       ELSIF "DB110_Interf_Program_M1".Status_IF[16].IF_is_on_1_Position AND "DB123_MH_IO_Signals".MH[16].IN.MH_Manual_Mode AND
           (#TempStationNo > 0 AND #TempStationNo < 101) THEN
           "DB619_State_MPart".ToolMa[#TmpMachineNumber].ToolNo := "DB941_Tool_alloc_manual_MH".MH[16].Alloc_stationTool[#TempStationNo];
       ELSE
           "DB619_State_MPart".ToolMa[#TmpMachineNumber].ToolNo := "DB940_Tool_alloc_automatic".Alloc_stationTool[#TempStationNo];
       END_IF;

       "DB619_State_MPart".ToolMa[#TmpMachineNumber].StationActive := True;
       "DB619_State_MPart".ToolMa[#TmpMachineNumber].StationNo := INT_TO_BYTE(#TempStationNo);
   END_IF;

   #TmpActToolNo := "DB619_State_MPart".ToolMa[#TmpMachineNumber].ToolNo;

   //-----------------------------------------------------------------
   // Check if tool no. between 1 and Amount tools if OK get data
   // ----------------------------------------------------------------
   IF (#TmpActToolNo > 0 AND
       #TmpActToolNo < "AmountTools") AND
      #IO_PartShotNoNew =  0 
    THEN
         #IO_PartShotNoNew:=  1;
         // Get tool values                                               
         "DB619_State_MPart".ToolMa[#TmpMachineNumber].Tool:= "DB930_Tools".Tool[#TmpActToolNo];
         // Get shot values; 
         IF (#TmpActToolNo > 0 AND
             #TmpActToolNo <= "AmountToolsDB")
         THEN
             "DB619_State_MPart".ShotMa[#TmpMachineNumber].Tool := "DB925_ShotData_1".Tool[#TmpActToolNo];

         ELSIF (#TmpActToolNo > "AmountToolsDB" AND #TmpActToolNo <= (2*"AmountToolsDB")) THEN
             "DB619_State_MPart".ShotMa[#TmpMachineNumber].Tool := "DB926_ShotData_2".Tool[#TmpActToolNo-"AmountToolsDB"];
         END_IF;

     ELSIF NOT (#TmpActToolNo > 0 AND #TmpActToolNo < "AmountToolsDB") THEN
         // Fault wrong tool no.    
         IF NOT #IO_Faults.FLT_WrongToolNumber AND
             "DB619_State_MPart".ToolMa[#TmpMachineNumber].StationActive AND
             NOT "DB619_State_MPart".ToolMa[#TmpMachineNumber].StationFinished THEN
               #IO_Faults.FLT_WrongToolNumber  := True;
               #IO_NewFault := True;
         END_IF;  
     END_IF;

   //-----------------------------------------------------------------------------------------
   // Check if new Tool is deselected 
   // ----------------------------------------------------------------------------------------
     IF NOT "DB619_State_MPart".ToolMa[#TmpMachineNumber].Tool.EnableTool AND
         "DB619_State_MPart".ToolMa[#TmpMachineNumber].StationActive THEN
         "DB619_State_MPart".ToolMa[#TmpMachineNumber].StationFinished := TRUE;
         "DB619_State_MPart".ToolMa[#TmpMachineNumber].ShotFound := FALSE;
         "DB619_State_MPart".ToolMa[#TmpMachineNumber].ToolNo := 0;
         "DB619_State_MPart".ToolMa[#TmpMachineNumber].PartShot := 0;
         "DB619_State_MPart".ShotMa[#TmpMachineNumber].ShotData.MH_No := 0;

         #IO_Faults.Reserve3 := TRUE;
   END_IF;


   //-----------------------------------------------------------------------------------------
   // Check if new partshot no. exist than get new MH no. and Shotvalues and set ShoFound 
   // ----------------------------------------------------------------------------------------
   IF #IO_PartShotNoNew <> "DB619_State_MPart".ToolMa[#TmpMachineNumber].PartShot AND
       "DB619_State_MPart".ToolMa[#TmpMachineNumber].StationActive
        THEN
            "DB619_State_MPart".ToolMa[#TmpMachineNumber].PartShot := #IO_PartShotNoNew;

         // Get mixinghead no. of selected part shot
            IF (#TmpActToolNo > 0 AND #TmpActToolNo < "AmountToolsDB") THEN
                #MH_No := "DB925_ShotData_1".Tool[#TmpActToolNo].Shot[#IO_PartShotNoNew].MHNo;
            ELSIF (#TmpActToolNo > "AmountToolsDB" AND #TmpActToolNo <= (2*"AmountToolsDB")) THEN
                #MH_No := "DB926_ShotData_2".Tool[#TmpActToolNo-"AmountToolsDB"].Shot[#IO_PartShotNoNew].MHNo;
            END_IF;

         "DB619_State_MPart".ShotMa[#TmpMachineNumber].ShotData.MH_No := INT_TO_BYTE(#MH_No);
             // Check mixinghead no. between 1 and 12
             IF #MH_No > 0 AND #MH_No < 13 THEN
                   // Mixinghead is connected at this machine
                   #MHNoShift := 1;
                   #MHNoBinary := SHL(IN :=  #MHNoShift, N := #MH_No -1);
                   #TmpMHatThisMachine := ("DB700_Machine".Machine[#TmpMachineNumber].MH_at_Machine AND #MHNoBinary) <> 0;
             ELSE
                   // Fault wrong mixinghead no. 
                 IF NOT  #IO_Faults.FLT_WrongMixingheadNumber AND "DB619_State_MPart".ToolMa[#TmpMachineNumber].StationActive THEN    // Must be wrong mixinghead no.                                                  
                     #IO_Faults.FLT_WrongMixingheadNumber := True;
                     #IO_Faults.FLT_WrongMixingheadNumber := False;
                     // #IO_NewFault := True;
                     //"DB619_State_MPart".ToolMa[#TmpMachineNumber].StationActive := FALSE;
                     //"DB619_State_MPart".ToolMa[#TmpMachineNumber].StationFinished := TRUE;
                 END_IF;
             END_IF;

   // Get shot values of current foamingcycle
             "DB619_State_MPart".ShotMa[#TmpMachineNumber].ShotData.ShotDisabled := "DB619_State_MPart".ShotMa[#TmpMachineNumber].Tool.Shot[#IO_PartShotNoNew].PartShotDisable;
             "DB619_State_MPart".ShotMa[#TmpMachineNumber].ShotData.CP_AfterShot := "DB619_State_MPart".ShotMa[#TmpMachineNumber].Tool.Shot[#IO_PartShotNoNew].CPMoveAfterShot;
             "DB619_State_MPart".ShotMa[#TmpMachineNumber].ShotData.Foamingtime := "DB619_State_MPart".ShotMa[#TmpMachineNumber].Tool.Shot[#IO_PartShotNoNew].FoamingTime;
             "DB619_State_MPart".ShotMa[#TmpMachineNumber].ShotData.PurgeMH_AfterShot := "DB619_State_MPart".ShotMa[#TmpMachineNumber].Tool.Shot[#IO_PartShotNoNew].PurgeMHAfterShot;

             "DB619_State_MPart".ShotMa[#TmpMachineNumber].ShotData.Flow[1] := "DB619_State_MPart".ShotMa[#TmpMachineNumber].Tool.Shot[#IO_PartShotNoNew].Flow[1];
             "DB619_State_MPart".ShotMa[#TmpMachineNumber].ShotData.Flow[2] := "DB619_State_MPart".ShotMa[#TmpMachineNumber].Tool.Shot[#IO_PartShotNoNew].Flow[2];
             "DB619_State_MPart".ShotMa[#TmpMachineNumber].ShotData.Flow[3] := "DB619_State_MPart".ShotMa[#TmpMachineNumber].Tool.Shot[#IO_PartShotNoNew].Flow[3];
             "DB619_State_MPart".ShotMa[#TmpMachineNumber].ShotData.Flow[4] := "DB619_State_MPart".ShotMa[#TmpMachineNumber].Tool.Shot[#IO_PartShotNoNew].Flow[4];
             "DB619_State_MPart".ShotMa[#TmpMachineNumber].ShotData.Flow[5] := "DB619_State_MPart".ShotMa[#TmpMachineNumber].Tool.Shot[#IO_PartShotNoNew].Flow[5];
             "DB619_State_MPart".ShotMa[#TmpMachineNumber].ShotData.Flow[6] := "DB619_State_MPart".ShotMa[#TmpMachineNumber].Tool.Shot[#IO_PartShotNoNew].Flow[6];
             "DB619_State_MPart".ShotMa[#TmpMachineNumber].ShotData.Pressure[1] := "DB619_State_MPart".ShotMa[#TmpMachineNumber].Tool.Shot[#IO_PartShotNoNew].Pressure[1];
             "DB619_State_MPart".ShotMa[#TmpMachineNumber].ShotData.Pressure[2] := "DB619_State_MPart".ShotMa[#TmpMachineNumber].Tool.Shot[#IO_PartShotNoNew].Pressure[2];
             "DB619_State_MPart".ShotMa[#TmpMachineNumber].ShotData.Pressure[3] := "DB619_State_MPart".ShotMa[#TmpMachineNumber].Tool.Shot[#IO_PartShotNoNew].Pressure[3];
             "DB619_State_MPart".ShotMa[#TmpMachineNumber].ShotData.Pressure[4] := "DB619_State_MPart".ShotMa[#TmpMachineNumber].Tool.Shot[#IO_PartShotNoNew].Pressure[4];
             "DB619_State_MPart".ShotMa[#TmpMachineNumber].ShotData.Pressure[5] := "DB619_State_MPart".ShotMa[#TmpMachineNumber].Tool.Shot[#IO_PartShotNoNew].Pressure[5];
             "DB619_State_MPart".ShotMa[#TmpMachineNumber].ShotData.Pressure[6] := "DB619_State_MPart".ShotMa[#TmpMachineNumber].Tool.Shot[#IO_PartShotNoNew].Pressure[6];

             "DB619_State_MPart".ShotMa[#TmpMachineNumber].ShotData."2PointAdjustment"[1] := "DB619_State_MPart".ShotMa[#TmpMachineNumber].Tool.Shot[#IO_PartShotNoNew]."2PoinMovement_Comp01";
             "DB619_State_MPart".ShotMa[#TmpMachineNumber].ShotData."2PointAdjustment"[2] := "DB619_State_MPart".ShotMa[#TmpMachineNumber].Tool.Shot[#IO_PartShotNoNew]."2PoinMovement_Comp02";
             "DB619_State_MPart".ShotMa[#TmpMachineNumber].ShotData."2PointAdjustment"[3] := "DB619_State_MPart".ShotMa[#TmpMachineNumber].Tool.Shot[#IO_PartShotNoNew]."2PoinMovement_Comp03";
             "DB619_State_MPart".ShotMa[#TmpMachineNumber].ShotData."2PointAdjustment"[4] := "DB619_State_MPart".ShotMa[#TmpMachineNumber].Tool.Shot[#IO_PartShotNoNew]."2PoinMovement_Comp04";
             "DB619_State_MPart".ShotMa[#TmpMachineNumber].ShotData."2PointAdjustment"[5] := "DB619_State_MPart".ShotMa[#TmpMachineNumber].Tool.Shot[#IO_PartShotNoNew]."2PoinMovement_Comp05";
             "DB619_State_MPart".ShotMa[#TmpMachineNumber].ShotData."2PointAdjustment"[6] := "DB619_State_MPart".ShotMa[#TmpMachineNumber].Tool.Shot[#IO_PartShotNoNew]."2PoinMovement_Comp06";

             "DB619_State_MPart".ShotMa[#TmpMachineNumber].ShotData.PartCounter := "DB619_State_MPart".ShotMa[#TmpMachineNumber].Tool.Shot[#IO_PartShotNoNew].PartCounter;


             "DB606_PV_Machine".Machine[#TmpMachineNumber].ShotTime.PV_SetV.Value := "DB619_State_MPart".ShotMa[#TmpMachineNumber].Tool.Shot[#IO_PartShotNoNew].FoamingTime;

   // Fault at tool is active      
   #IO_FaultAtStation := #IO_Faults.FLT_WrongToolNumber       OR
                         #IO_Faults.FLT_WrongMixingheadNumber OR
                         #IO_Faults.FLT_NewNoTooEarly;

   // Set shot found if tool is enabled                      
                         IF "DB619_State_MPart".ToolMa[#TmpMachineNumber].StationActive  AND NOT
                                              #IO_FaultAtStation  AND
                                              #IN_EnableTool      AND
                                              #TmpMHatThisMachine AND
                                              "DB619_State_MPart".ToolMa[#TmpMachineNumber].Tool.EnableTool
      THEN            
          "DB619_State_MPart".ToolMa[#TmpMachineNumber].ShotFound := True;
      ELSE       
          "DB619_State_MPart".ToolMa[#TmpMachineNumber].ShotFound := FALSE;
      END_IF;
    END_IF;

   //------------------------------------------------------------------------------------------
   // New Partshot no. -> Shotend, Shotbreak, next shot at this machine
   // -----------------------------------------------------------------------------------------
    IF  ("DB619_State_MPart".ToolMa[#TmpMachineNumber].StationActive AND NOT
        "DB619_State_MPart".ToolMa[#TmpMachineNumber].ShotFound)     OR
        "DB619_State_MPart".Cycle[#TmpMachineNumber].PulsShotend
       THEN  
           IF "DB619_State_MPart".ToolMa[#TmpMachineNumber].PartShot <= BYTE_TO_INT("DB619_State_MPart".ToolMa[#TmpMachineNumber].Tool.PartShot_Amount) THEN
               #IO_PartShotNoNew := "DB619_State_MPart".ToolMa[#TmpMachineNumber].PartShot + 1;
               "DB619_State_MPart".ToolMa[#TmpMachineNumber].ShotFound := FALSE;
           END_IF;

       END_IF;

       // Station finished: shots done; cycle stopped; fault level 1; station no. = 0
       IF "DB619_State_MPart".ToolMa[#TmpMachineNumber].PartShot > BYTE_TO_INT("DB619_State_MPart".ToolMa[#TmpMachineNumber].Tool.PartShot_Amount) OR
          "DB009_Faults".Fault_State_Grp_1_M1                 OR
          "DB619_State_MPart".ToolMa[#TmpMachineNumber].StopCycle
       THEN
           "DB619_State_MPart".ToolMa[#TmpMachineNumber].StationFinished := TRUE;
           "DB619_State_MPart".ToolMa[#TmpMachineNumber].ShotFound := FALSE;
           "DB619_State_MPart".ToolMa[#TmpMachineNumber].ToolNo := 0;
           "DB619_State_MPart".ToolMa[#TmpMachineNumber].PartShot := 0;
           "DB619_State_MPart".ShotMa[#TmpMachineNumber].ShotData.MH_No := 0;
       END_IF;

       IF  #IO_Faults.FLT_WrongToolNumber       OR
           #IO_Faults.FLT_WrongMixingheadNumber OR
           #IO_Faults.FLT_NewNoTooEarly         OR
           #IO_Faults.Reserve3
         THEN
           #IO_FaultLevel_1 := TRUE;
       END_IF;
END_FUNCTION_BLOCK

FUNCTION_BLOCK "FB1931_ToolAllocationList"   // FB1931, SCL
{ S7_Optimized_Access := 'TRUE' }
VERSION : 0.1
   VAR
      Alloc_stationTool : Array[0..30] of Int;
      SaveSortProgs : Array[0..20] of Int;
   END_VAR
   VAR_TEMP
      j : Int;
      i : Int;
      z : Int;
      TiLoop : Int;
      TiLoopSave : Int;
      TiLoopMH : Int;
      Ti_alloc_list : Int;
      Amount_tools : Int;
      MH_No_hand_allocation : Int;
      Offset_SavedProgsList : Int;
      Offset_AllocateList : Int;
      LimitSavedProgList : Int;
      Amount_Saved_tools : Int;
      tool_okay : Bool;
   END_VAR
   // Alloc_stationTool[0] := 0;
   // Alloc_stationTool[1] := 0;
   // Alloc_stationTool[2] := 0;
   // Alloc_stationTool[3] := 0;
   // Alloc_stationTool[4] := 0;
   // Alloc_stationTool[5] := 0;
   // Alloc_stationTool[6] := 0;
   // Alloc_stationTool[7] := 0;
   // Alloc_stationTool[8] := 0;
   // Alloc_stationTool[9] := 0;
   // Alloc_stationTool[10] := 0;
   // Alloc_stationTool[11] := 0;
   // Alloc_stationTool[12] := 0;
   // Alloc_stationTool[13] := 0;
   // Alloc_stationTool[14] := 0;
   // Alloc_stationTool[15] := 0;
   // Alloc_stationTool[16] := 0;
   // Alloc_stationTool[17] := 0;
   // Alloc_stationTool[18] := 0;
   // Alloc_stationTool[19] := 0;
   // Alloc_stationTool[20] := 0;
   // Alloc_stationTool[21] := 0;
   // Alloc_stationTool[22] := 0;
   // Alloc_stationTool[23] := 0;
   // Alloc_stationTool[24] := 0;
   // Alloc_stationTool[25] := 0;
   // Alloc_stationTool[26] := 0;
   // Alloc_stationTool[27] := 0;
   // Alloc_stationTool[28] := 0;
   // Alloc_stationTool[29] := 0;
   // Alloc_stationTool[30] := 0;
BEGIN
   // Limit values

   "DB939_Tool_alloc_HMI".Selected_prog := LIMIT(MN := 1, IN := "DB939_Tool_alloc_HMI".Selected_prog, MX := 30);
   "DB939_Tool_alloc_HMI".Selected_SavedProg := LIMIT(MN := 0, IN := "DB939_Tool_alloc_HMI".Selected_SavedProg, MX := 20);
   "DB939_Tool_alloc_HMI".Limit_allocation_list := LIMIT(MN := 1, IN := "DB939_Tool_alloc_HMI".Limit_allocation_list, MX := 30);

   FOR #TiLoop := 0 TO 30 DO
       "DB939_Tool_alloc_HMI".Alloc_stationTool[#TiLoop] := LIMIT(MN := 0, IN := "DB939_Tool_alloc_HMI".Alloc_stationTool[#TiLoop], MX := "AmountTools");
   END_FOR;

   REGION Select manual/auto
       // Switch for choosing manual or automatic allocation on the Screen "ProgramAllocation"  
       IF "DB939_Tool_alloc_HMI".Select_hand_automatic_alloc = TRUE THEN
           "DB939_Tool_alloc_HMI".Tool_allocation_automatic := FALSE;
           "DB939_Tool_alloc_HMI".Tool_allocation_manual := TRUE;
       ELSE
           "DB939_Tool_alloc_HMI".Tool_allocation_automatic := TRUE;
           "DB939_Tool_alloc_HMI".Tool_allocation_manual := FALSE;
       END_IF;
   END_REGION

   // Current selected mixing head number for Hand allocation
   #MH_No_hand_allocation := "DB939_Tool_alloc_HMI".MH_No_selected;

   REGION Visibility MH arrows 
       // Visibility of arrow for decreasing Mixing head number
       IF "DB939_Tool_alloc_HMI".Tool_allocation_manual = TRUE AND #MH_No_hand_allocation > 1 THEN
           "DB939_Tool_alloc_HMI".MH_Nr_decrease_visible := TRUE;
       ELSE
           "DB939_Tool_alloc_HMI".MH_Nr_decrease_visible := FALSE;
       END_IF;

       // Visibility of arrow for increasing Mixing head number
       IF "DB939_Tool_alloc_HMI".Tool_allocation_manual = TRUE AND #MH_No_hand_allocation < "DB790_PlantParameter".AmountMH THEN
           "DB939_Tool_alloc_HMI".MH_Nr_increase_visible := TRUE;
       ELSE
           "DB939_Tool_alloc_HMI".MH_Nr_increase_visible := FALSE;
       END_IF;
   END_REGION

   REGION Page AllocationList
       // Depending on amound of manual programs limit list and pages
       IF "DB704_MH_Value".Mixinghead[#MH_No_hand_allocation].With99program = FALSE AND "DB939_Tool_alloc_HMI".Tool_allocation_automatic = FALSE THEN
           "DB939_Tool_alloc_HMI".Limit_allocation_page := 1;
           "DB939_Tool_alloc_HMI".Limit_allocation_list := 9;
       ELSIF "DB704_MH_Value".Mixinghead[#MH_No_hand_allocation].With99program = TRUE AND "DB939_Tool_alloc_HMI".Tool_allocation_automatic = FALSE THEN
           "DB939_Tool_alloc_HMI".Limit_allocation_page := 4;
           IF "DB939_Tool_alloc_HMI".AllocList_page >= 4 THEN
               "DB939_Tool_alloc_HMI".Limit_allocation_list := 9;
           ELSE
               "DB939_Tool_alloc_HMI".Limit_allocation_list := 30;
           END_IF;
       ELSIF "DB939_Tool_alloc_HMI".Tool_allocation_automatic = TRUE THEN
         //Depending on the amount of the stationsnumber   
           "DB939_Tool_alloc_HMI".Limit_allocation_page := (("DB790_PlantParameter".AmountToolStation -1 ) / (30))+1;
           IF "DB939_Tool_alloc_HMI".AllocList_page = "DB939_Tool_alloc_HMI".Limit_allocation_page  AND ("DB790_PlantParameter".AmountToolStation MOD 30) <> 0 THEN
               "DB939_Tool_alloc_HMI".Limit_allocation_list := ("DB790_PlantParameter".AmountToolStation MOD 30);
           ELSE
               "DB939_Tool_alloc_HMI".Limit_allocation_list := 30;
           END_IF;
       ELSE   
           "DB939_Tool_alloc_HMI".Limit_allocation_page := 7;
           "DB939_Tool_alloc_HMI".Limit_allocation_list := 30;
       END_IF;

       IF "DB939_Tool_alloc_HMI".AllocList_increase THEN
           "DB939_Tool_alloc_HMI".AllocList_page := "DB939_Tool_alloc_HMI".AllocList_page + 1;
           "DB939_Tool_alloc_HMI".AllocList_increase := False;
       ELSIF "DB939_Tool_alloc_HMI".AllocList_decrease THEN
           "DB939_Tool_alloc_HMI".AllocList_page := "DB939_Tool_alloc_HMI".AllocList_page - 1;
           "DB939_Tool_alloc_HMI".AllocList_decrease := False;
       END_IF;
       // Limit
       "DB939_Tool_alloc_HMI".AllocList_page := LIMIT(MN := 1, IN := "DB939_Tool_alloc_HMI".AllocList_page, MX := "DB939_Tool_alloc_HMI".Limit_allocation_page);
       // Create offset
       #Offset_AllocateList := ("DB939_Tool_alloc_HMI".AllocList_page - 1) * 30;
   END_REGION

   REGION Useable Alloc arrows
    // This part is used for if you can alloc the programm to the allocaationlist by yourself 
    // or automatically by the inferface
       IF "DB939_Tool_alloc_HMI".Tool_allocation_automatic = TRUE AND "DB790_PlantParameter".Bit.ProgrammNofromInterface = TRUE THEN
           IF  ("DB790_PlantParameter".AmountMouldCarrier MOD 30) <> 0 THEN
               IF "DB939_Tool_alloc_HMI".AllocList_page = ((("DB790_PlantParameter".AmountMouldCarrier - 1) / 30)+1) THEN
                    "DB939_Tool_alloc_HMI".Operability_selected_line := ("DB790_PlantParameter".AmountMouldCarrier MOD 30);
                ELSIF   "DB939_Tool_alloc_HMI".AllocList_page < ((("DB790_PlantParameter".AmountMouldCarrier - 1) / 30)+1) THEN
                   "DB939_Tool_alloc_HMI".Operability_selected_line := 30;
                ELSE
                   "DB939_Tool_alloc_HMI".Operability_selected_line := 0;
               END_IF;
           ELSE
               IF "DB939_Tool_alloc_HMI".AllocList_page <= ((("DB790_PlantParameter".AmountMouldCarrier - 1) / 30)+1) THEN
                    "DB939_Tool_alloc_HMI".Operability_selected_line := 30;
               ELSE
                   "DB939_Tool_alloc_HMI".Operability_selected_line := 0;
               END_IF;
           END_IF;
       ELSE 
           "DB939_Tool_alloc_HMI".Operability_selected_line := 0;
       END_IF;

       IF "DB939_Tool_alloc_HMI".Selected_prog <= "DB939_Tool_alloc_HMI".Operability_selected_line THEN
           "DB939_Tool_alloc_HMI".Selected_prog := 0;
       END_IF;
   END_REGION
   REGION Visibility Alloc arrows
       IF "DB939_Tool_alloc_HMI".AllocList_page < "DB939_Tool_alloc_HMI".Limit_allocation_page THEN
           "DB939_Tool_alloc_HMI".AllocList_increase_visible := TRUE;
       ELSE    
           "DB939_Tool_alloc_HMI".AllocList_increase_visible := FALSE;
       END_IF;

       IF "DB939_Tool_alloc_HMI".AllocList_page > 1 THEN
           "DB939_Tool_alloc_HMI".AllocList_decrease_visible := TRUE;
       ELSE
           "DB939_Tool_alloc_HMI".AllocList_decrease_visible := FALSE;
       END_IF;
   END_REGION

   REGION Page SavedProgsList
       // Depending on the saved tools. Limit saved list
       #Amount_Saved_tools := 0;
       FOR #TiLoop := 1 TO "AmountTools" DO
           IF "DB933_SaveSortProgs".SaveSortTool[#TiLoop] <> 0 THEN
               #Amount_Saved_tools := #Amount_Saved_tools + 1;
           END_IF;
       END_FOR;
       IF #Amount_Saved_tools > 0 THEN
           #LimitSavedProgList := ((#Amount_Saved_tools - 1) / 20) + 1;
       ELSE
           #LimitSavedProgList := 1;
       END_IF;


       IF "DB939_Tool_alloc_HMI".SavedProgs_increase THEN
           "DB939_Tool_alloc_HMI".SavedProgs_page := "DB939_Tool_alloc_HMI".SavedProgs_page + 1;
           "DB939_Tool_alloc_HMI".SavedProgs_increase := False;
       ELSIF "DB939_Tool_alloc_HMI".SavedProgs_decrease THEN
           "DB939_Tool_alloc_HMI".SavedProgs_page := "DB939_Tool_alloc_HMI".SavedProgs_page - 1;
           "DB939_Tool_alloc_HMI".SavedProgs_decrease := False;
       END_IF;
       // Limit
       "DB939_Tool_alloc_HMI".SavedProgs_page := LIMIT(MN := 1, IN := "DB939_Tool_alloc_HMI".SavedProgs_page, MX := #LimitSavedProgList);
       // Create offset
       #Offset_SavedProgsList := ("DB939_Tool_alloc_HMI".SavedProgs_page - 1) * 20;
   END_REGION

   REGION Visibility SavedProgList arrows
       IF "DB939_Tool_alloc_HMI".SavedProgs_page < #LimitSavedProgList THEN
           "DB939_Tool_alloc_HMI".SavedProgs_increase_visible := TRUE;
       ELSE
           "DB939_Tool_alloc_HMI".SavedProgs_increase_visible := FALSE;
       END_IF;

       IF "DB939_Tool_alloc_HMI".SavedProgs_page > 1 THEN
           "DB939_Tool_alloc_HMI".SavedProgs_decrease_visible := TRUE;
       ELSE
           "DB939_Tool_alloc_HMI".SavedProgs_decrease_visible := FALSE;
       END_IF;
   END_REGION

   REGION Clear SavedProgsList
       FOR #z := 0 TO "AmountTools" DO
           // Clear list
           "DB933_SaveSortProgs".SaveSortTool[#z] := 0;
       END_FOR;
   END_REGION

   REGION Create SavedProgsList
       // Check if part shots available or not for allocation list
       #j := 1;
       FOR #TiLoop := 1 TO "AmountTools" DO
           IF "DB930_Tools".Tool[#TiLoop].PartShot_Amount <> 0 THEN
               "DB933_SaveSortProgs".SaveSortTool[#j] := #TiLoop;
               #j := #j + 1;
           END_IF;
       END_FOR;
   END_REGION

   REGION Copy Part of list savedprogslist to actual HMI
       FOR #TiLoop := 1 TO 20 DO
           "DB939_Tool_alloc_HMI".SaveSortProgs[#TiLoop] := "DB933_SaveSortProgs".SaveSortTool[#TiLoop + #Offset_SavedProgsList];
       END_FOR;
   END_REGION

   REGION Delete selected tool allocation
       IF "DB939_Tool_alloc_HMI".Delete_selected_tool <> 0 THEN
           "DB939_Tool_alloc_HMI".Alloc_stationTool["DB939_Tool_alloc_HMI".Delete_selected_tool] := 0;
           "DB939_Tool_alloc_HMI".Delete_selected_tool := 0;
       END_IF;
   END_REGION

   REGION Delete selected tool from Mould Editor in all allocation lists
       IF "DB939_Tool_alloc_HMI"."Delete_tool_in _all_allocations" AND "DB_MouldEditor_HMI".uData.sStatusBits.xFaultDeleteProgram THEN
           // search tool in automatic allocation list
           FOR #TiLoop := 1 TO "InterfaceVisu".AmountAlloactionAutomatic DO
               IF "DB940_Tool_alloc_automatic".Alloc_stationTool[#TiLoop] = "DB_MouldEditor_HMI".uData.sSelected.iTool THEN
                   "DB940_Tool_alloc_automatic".Alloc_stationTool[#TiLoop] := 0;
               END_IF;
           END_FOR;
           // search tool in all manual allocation lists
           FOR #TiLoopMH := 1 TO "DB790_PlantParameter".AmountMH DO
               IF "DB704_MH_Value".Mixinghead[#TiLoopMH].With99program THEN
                   #Ti_alloc_list := 99;
               ELSE
                   #Ti_alloc_list := 9;
               END_IF;

               FOR #TiLoop := 1 TO #Ti_alloc_list DO
                   IF "DB941_Tool_alloc_manual_MH".MH[#TiLoopMH].Alloc_stationTool[#TiLoop] = "DB_MouldEditor_HMI".uData.sSelected.iTool THEN
                       "DB941_Tool_alloc_manual_MH".MH[#TiLoopMH].Alloc_stationTool[#TiLoop] := 0;
                   END_IF;
               END_FOR;
           END_FOR;
           // reset bits to delete and for PopUp
           "DB939_Tool_alloc_HMI"."Delete_tool_in _all_allocations" := FALSE;
           "DB_MouldEditor_HMI".uData.sStatusBits.xFaultDeleteProgram := FALSE;
           "DB_MouldEditor_HMI".uData.sStatusBits.xDeleteProgram := TRUE; // <-- delete tool
       END_IF;
   END_REGION

   REGION assign saved tool to selected tool    
       IF "DB939_Tool_alloc_HMI".Selected_SavedProg <> 0 THEN
           // If no programm is allocated set new programm
           IF "DB939_Tool_alloc_HMI".Alloc_stationTool["DB939_Tool_alloc_HMI".Selected_prog] = 0 THEN
               "DB939_Tool_alloc_HMI".Alloc_stationTool["DB939_Tool_alloc_HMI".Selected_prog] := "DB933_SaveSortProgs".SaveSortTool["DB939_Tool_alloc_HMI".Selected_SavedProg + #Offset_SavedProgsList];
               "DB939_Tool_alloc_HMI".Selected_SavedProg := 0;
               "DB939_Tool_alloc_HMI".Overwrite_not_allowed := FALSE;
           ELSIF "DB939_Tool_alloc_HMI".Alloc_stationTool["DB939_Tool_alloc_HMI".Selected_prog] = "DB933_SaveSortProgs".SaveSortTool["DB939_Tool_alloc_HMI".Selected_SavedProg + #Offset_SavedProgsList] THEN
               "DB939_Tool_alloc_HMI".Selected_SavedProg := 0;
           ELSE
               "DB939_Tool_alloc_HMI".Overwrite_not_allowed := TRUE;
               IF "DB939_Tool_alloc_HMI".Overwrite_selected_tool = TRUE THEN
                   "DB939_Tool_alloc_HMI".Alloc_stationTool["DB939_Tool_alloc_HMI".Selected_prog] := "DB933_SaveSortProgs".SaveSortTool["DB939_Tool_alloc_HMI".Selected_SavedProg + #Offset_SavedProgsList];
                   "DB939_Tool_alloc_HMI".Selected_SavedProg := 0;
                   "DB939_Tool_alloc_HMI".Overwrite_not_allowed := FALSE;
                   "DB939_Tool_alloc_HMI".Overwrite_selected_tool := FALSE;
               END_IF;
           END_IF;
       ELSE    
           "DB939_Tool_alloc_HMI".Overwrite_not_allowed := FALSE;
       END_IF;
   END_REGION

   REGION Allocationlist number changed
       // If any allocation list no changed, store it to the right DB
       FOR #TiLoop := 1 TO 30 DO
           IF "DB939_Tool_alloc_HMI".Alloc_stationTool[#TiLoop] <> #Alloc_stationTool[#TiLoop] THEN
               IF "DB939_Tool_alloc_HMI".Tool_allocation_automatic = TRUE THEN
                   "DB940_Tool_alloc_automatic".Alloc_stationTool[#TiLoop + #Offset_AllocateList] := "DB939_Tool_alloc_HMI".Alloc_stationTool[#TiLoop];
               ELSE
                   "DB941_Tool_alloc_manual_MH".MH["DB939_Tool_alloc_HMI".MH_No_selected].Alloc_stationTool[#TiLoop + #Offset_AllocateList] := "DB939_Tool_alloc_HMI".Alloc_stationTool[#TiLoop];
               END_IF;
           END_IF;
       END_FOR;
   END_REGION

   REGION Copy Part of allocat list to actual HMI


       FOR #TiLoop := 1 TO 30 DO
           IF "DB939_Tool_alloc_HMI".Tool_allocation_automatic = TRUE THEN
               "DB939_Tool_alloc_HMI".Alloc_stationTool[#TiLoop] := "DB940_Tool_alloc_automatic".Alloc_stationTool[#TiLoop + #Offset_AllocateList];
           ELSE
               "DB939_Tool_alloc_HMI".Alloc_stationTool[#TiLoop] := "DB941_Tool_alloc_manual_MH".MH["DB939_Tool_alloc_HMI".MH_No_selected].Alloc_stationTool[#TiLoop + #Offset_AllocateList];
           END_IF;
           // Depending on BCD switch load 9 or 30 (99) programs in the list
           IF ("DB704_MH_Value".Mixinghead[#MH_No_hand_allocation].With99program = FALSE AND "DB939_Tool_alloc_HMI".Tool_allocation_automatic = FALSE AND #TiLoop >= 9)
               OR ("DB704_MH_Value".Mixinghead[#MH_No_hand_allocation].With99program = TRUE AND "DB939_Tool_alloc_HMI".Tool_allocation_automatic = FALSE AND #TiLoop >= 9 AND "DB939_Tool_alloc_HMI".AllocList_page >= 4) THEN
               EXIT;
           END_IF;
       END_FOR;
   END_REGION

   REGION Copy tool names to actual HMI lists
       FOR #TiLoop := 1 TO 30 DO
           IF "DB939_Tool_alloc_HMI".Alloc_stationTool[#TiLoop] <= "AmountTools" THEN
               "DB939_Tool_alloc_HMI".Alloc_tool_name[#TiLoop] := "DB930_Tools".Tool["DB939_Tool_alloc_HMI".Alloc_stationTool[#TiLoop]].tool_name;
           END_IF;
       END_FOR;
       FOR #TiLoop := 1 TO 20 DO
           "DB939_Tool_alloc_HMI".SaveSortProg_name[#TiLoop] := "DB930_Tools".Tool["DB939_Tool_alloc_HMI".SaveSortProgs[#TiLoop]].tool_name;
       END_FOR;
   END_REGION

   REGION Wrong tool allocated
       // Delete tool from all lists if it's not in the saved progs list
       "DB939_Tool_alloc_HMI".Tool_not_exist := FALSE; // <-- no pop up
       FOR #TiLoop := 1 TO "AmountAllocationAutomatic" DO
           #tool_okay := FALSE;
           FOR #TiLoopSave := 1 TO "AmountTools" DO
               IF "DB940_Tool_alloc_automatic".Alloc_stationTool[#TiLoop] = "DB933_SaveSortProgs".SaveSortTool[#TiLoopSave] THEN
                   #tool_okay := TRUE;
                   EXIT;
               // Stop loop at first "0" in SavedToolsList or if Loop number is higher then the allocated tool number    
               ELSIF "DB933_SaveSortProgs".SaveSortTool[#TiLoopSave] = 0 OR #TiLoopSave > "DB940_Tool_alloc_automatic".Alloc_stationTool[#TiLoop] THEN
                   EXIT;
               END_IF;
           END_FOR;
           IF #tool_okay = FALSE THEN
               "DB940_Tool_alloc_automatic".Alloc_stationTool[#TiLoop] := 0;
               #tool_okay := FALSE;
           END_IF;
       END_FOR;
       // Manual allocation list
       FOR #TiLoopMH := 1 TO "DB790_PlantParameter".AmountMH DO
           FOR #TiLoop := 1 TO 120 DO // <-- all tools also if only 9 or 99 possible
               FOR #TiLoopSave := 1 TO "AmountTools" DO
                   #tool_okay := FALSE;
                   IF "DB941_Tool_alloc_manual_MH".MH[#TiLoopMH].Alloc_stationTool[#TiLoop] = "DB933_SaveSortProgs".SaveSortTool[#TiLoopSave] THEN
                       #tool_okay := TRUE;
                       EXIT;
                       // Stop loop at first "0" in SavedToolsList or if Loop number is higher then the allocated tool number    
                   ELSIF "DB933_SaveSortProgs".SaveSortTool[#TiLoopSave] = 0 OR #TiLoopSave > "DB941_Tool_alloc_manual_MH".MH[#TiLoopMH].Alloc_stationTool[#TiLoop] THEN
                       EXIT;
                   END_IF;
               END_FOR;
               IF #tool_okay = FALSE THEN
                   "DB941_Tool_alloc_manual_MH".MH[#TiLoopMH].Alloc_stationTool[#TiLoop] := 0;
                   #tool_okay := FALSE;
               END_IF;
           END_FOR;
       END_FOR;
   END_REGION

   REGION Save DB
       FOR #TiLoop := 1 TO 30 DO
           #Alloc_stationTool[#TiLoop] := "DB939_Tool_alloc_HMI".Alloc_stationTool[#TiLoop];
       END_FOR;
   END_REGION
END_FUNCTION_BLOCK

FUNCTION "GWK_PB_TecoCS(CW)e" : Void   // FC1, SCL
TITLE = GWK_PB_TecoEP
{ S7_Optimized_Access := 'FALSE' }
AUTHOR : SCDE
FAMILY : GWK
NAME : PBcomEP
VERSION : 1.3
// TecoCS/CW
// GWK ProfiBus Kommunikation Einfaches Protokoll mit Systemfunktionen SFC 14 SFC 15 und SFC 21 (Löschung)
// 
//  KNOW_HOW_PROTECT
// ////////
//  Änderungen
// 
//   
//     V1.3:
//     Startwertinitialisierung fällt weg
//     
//     V1.2:
//     Istwerttelegramm wird nur in DB kopiert bei fehlerfreier Abarbeitung SFC 14 und SL_akt
//     
//     V1.1: 
//     zusätzliche Sicht "BYTE" für die Sende- und Empfangsdaten eingefügt, da auf einem kundenseitigen S7-400 System die SFC 14/15 einen 8092 Fehler zurück meldeten 
//     (ANY POINTER liegt nicht im BYTE Format vor). Nun erstellt der Kompiler einen Byte-Formatierten Zeiger.
//   
//     V1.0: 
//     Ursprungsversion
// 
// ////////
//  Bausteinparameter
   VAR_INPUT
      IN_With_tempering_unit : Bool;   // Mouldcarrier has an tempering unit
      IN_Flag_alarm : Bool;   // Pulseflag for alarm list
      IN_Adr : Hw_Any;   // Hardwarekonfig
      IN_Sl_Akt : Bool;   // Slave aktiv; 1 = Abarbeitung SFC14/15; 0 = keine Abarbeitung SFC14/15, Telegramme löschen
      IN_TL_KomF : Bool;   // 1 = Telegramme löschen bei SFC 14 Kommunikationsfehler; 0 = Telegramme behalten
      IN_On : Bool;   // On/Off
      IN_Release : Bool;   // Release
      IN_Weekendmode : Bool;   // Temperaturabsenkung aktivieren
      IN_Fault_quit : Bool;   // Quit faults
      IN_Fuse : Bool;   // Fault fuse
      IN_Setvalue : Int;   // Temperature setvalue
      IN_Setvalue_weekend : Int;   // Temperature setvalue weekend
      IN_Actvalue_tool : Real;   // Actual temperature tool
   END_VAR
   VAR_IN_OUT
      RetVal_SFC14 : Word;   // Rückgabewert Systemfunktion SFC 14
      RetVal_SFC15 : Word;   // Rückgabewert Systemfunktion SFC 15
      PBData : "PB_TecoCS(CW)e_SW-IW";
      Sicht_word AT PBData : Array[0..11] of Word;
      Sicht_Byte AT PBData : Array[0..23] of Byte;
      Sicht_bool AT PBData : Array[0..15] of Bool;
      State : "UDT_State_GWK";
   END_VAR
   VAR_TEMP
      Sendedaten : Array[0..5] of Word;
      Sendedaten_BYTE AT Sendedaten : Array[0..11] of Byte;   // V1.1
      Empfangsdaten : Array[0..5] of Word;
      Empfangsdaten_BYTE AT Empfangsdaten : Array[0..11] of Byte;   // V1.1
      index : Int;
      State_index : Int;
      Temp_state : Word;
   END_VAR
BEGIN
   IF #IN_With_tempering_unit THEN
     // Sendedaten aus DB in den Temp. Puffer kopieren

     FOR #index := 0 TO 5 DO
       #Sendedaten[#index] := #Sicht_word[#index];
     END_FOR;

     // ProfiNet daten lesen
     IF #IN_Sl_Akt THEN
       #RetVal_SFC14 := INT_TO_WORD(DPRD_DAT(LADDR := #IN_Adr, RECORD => #Empfangsdaten_BYTE));
     ELSE
       #RetVal_SFC14 := 0;
     END_IF;

     // Sollwertvorgabe
     IF #IN_Weekendmode = true THEN
       #PBData.SW.T1W2 := #IN_Setvalue_weekend;
     ELSE
       #PBData.SW.T1W2 := #IN_Setvalue;
     END_IF;

     // Limit (relative to setpoint)
     #PBData.SW.T1W3 := 100;
     // Max. flow line temperature
     #PBData.SW.T1W4 := 1000;

     // Switch on
     #PBData.SW.W1.Bit0 := #IN_On AND #IN_Release;
     // Ext. Sensor
     #PBData.SW.W1.Bit1 := 0;
     // Normal operation
     #PBData.SW.W1.Bit2 := 1;
     // Standby operation
     #PBData.SW.W1.Bit3 := 0;
     // Leak stop operation
     #PBData.SW.W1.Bit4 := 0;
     // Mould draining
     #PBData.SW.W1.Bit5 := 0;
     // Cool down unit and switch off
     #PBData.SW.W1.Bit6 := 0;
     // Monitoring limit value
     #PBData.SW.W1.Bit7 := 0;
     REGION #State for HMI
       // ON
       #State.on := #PBData.IW.T1_W2.Bit2;
       // Fault
       IF #Sicht_word[6] > 1 THEN
         #State.Fault := TRUE;
       ELSE
         #State.Fault := FALSE;
       END_IF;
       // Weekend mode
       #State.Weekend_mode := #IN_Weekendmode;
       // Set value
       #State.Set_value_tempering_unit := #PBData.SW.T1W2;
       // Act value
       #State.Act_value_tempering_unit := INT_TO_REAL((#PBData.IW.T1_W3)) / real#10.0;
       // Act value tool
       #State.Act_value_tool := REAL_TO_INT(#IN_Actvalue_tool);
     END_REGION

     REGION #Generate state
       // Each second the new alarm number is showed on the TP
       IF #IN_Flag_alarm THEN

         IF #PBData.IW.T1_W1.Bit0 AND #State.Fault = FALSE AND #State.Fault_index = 0 AND #State.Fault_state <> 1 THEN
           #State.Fault_state := 1;
           #State.Fault_index := #State.Fault_index + 1;
         ELSIF #PBData.IW.T1_W1.Bit1 AND #State.Fault_index >= 0 AND #State.Fault_index <= 1 AND #State.Fault_state <> 2 THEN
           #State.Fault_state := 2;
           #State.Fault_index := #State.Fault_index + 1;
         ELSIF #PBData.IW.T1_W1.Bit2 AND #State.Fault_index >= 0 AND #State.Fault_index <= 2 AND #State.Fault_state <> 3 THEN
           #State.Fault_state := 3;
           #State.Fault_index := #State.Fault_index + 1;
         ELSIF #PBData.IW.T1_W1.Bit3 AND #State.Fault_index >= 0 AND #State.Fault_index <= 3 AND #State.Fault_state <> 4 THEN
           #State.Fault_state := 4;
           #State.Fault_index := #State.Fault_index + 1;
         ELSIF #PBData.IW.T1_W1.Bit4 AND #State.Fault_index >= 0 AND #State.Fault_index <= 4 AND #State.Fault_state <> 5 THEN
           #State.Fault_state := 5;
           #State.Fault_index := #State.Fault_index + 1;
         ELSIF #PBData.IW.T1_W1.Bit5 AND #State.Fault_index >= 0 AND #State.Fault_index <= 5 AND #State.Fault_state <> 6 THEN
           #State.Fault_state := 6;
           #State.Fault_index := #State.Fault_index + 1;
         ELSIF #PBData.IW.T1_W1.Bit6 AND #State.Fault_index >= 0 AND #State.Fault_index <= 6 AND #State.Fault_state <> 7 THEN
           #State.Fault_state := 7;
           #State.Fault_index := #State.Fault_index + 1;
         ELSIF #PBData.IW.T1_W1.Bit7 AND #State.Fault_index >= 0 AND #State.Fault_index <= 7 AND #State.Fault_state <> 8 THEN
           #State.Fault_state := 8;
           #State.Fault_index := #State.Fault_index + 1;
         ELSIF #PBData.IW.T1_W1.Bit8 AND #State.Fault_index >= 0 AND #State.Fault_index <= 8 AND #State.Fault_state <> 9 THEN
           #State.Fault_state := 9;
           #State.Fault_index := #State.Fault_index + 1;
         ELSIF #PBData.IW.T1_W1.Bit9 AND #State.Fault_index >= 0 AND #State.Fault_index <= 9 AND #State.Fault_state <> 10 THEN
           #State.Fault_state := 10;
           #State.Fault_index := #State.Fault_index + 1;
         ELSIF #PBData.IW.T1_W1.Bit10 AND #State.Fault_index >= 0 AND #State.Fault_index <= 10 AND #State.Fault_state <> 11 THEN
           #State.Fault_state := 11;
           #State.Fault_index := #State.Fault_index + 1;
         ELSIF #PBData.IW.T1_W1.Bit11 AND #State.Fault_index >= 0 AND #State.Fault_index <= 11 AND #State.Fault_state <> 12 THEN
           #State.Fault_state := 12;
           #State.Fault_index := #State.Fault_index + 1;
         ELSIF #PBData.IW.T1_W1.Bit12 AND #State.Fault_index >= 0 AND #State.Fault_index <= 12 AND #State.Fault_state <> 13 THEN
           #State.Fault_state := 13;
           #State.Fault_index := #State.Fault_index + 1;
         ELSIF #PBData.IW.T1_W1.Bit13 AND #State.Fault_index >= 0 AND #State.Fault_index <= 13 AND #State.Fault_state <> 14 THEN
           #State.Fault_state := 14;
           #State.Fault_index := #State.Fault_index + 1;
         ELSIF #PBData.IW.T1_W1.Bit14 AND #State.Fault_index >= 0 AND #State.Fault_index <= 14 AND #State.Fault_state <> 15 THEN
           #State.Fault_state := 15;
           #State.Fault_index := #State.Fault_index + 1;
         ELSIF #PBData.IW.T1_W1.Bit15 AND #State.Fault_index >= 0 AND #State.Fault_index <= 15 AND #State.Fault_state <> 16 THEN
           #State.Fault_state := 16;
           #State.Fault_index := #State.Fault_index + 1;

         ELSIF #PBData.IW.T1_W2.Bit0 = false AND #State.Fault_index >= 0 AND #State.Fault_index <= 16 AND #State.Fault_state <> 17 THEN
           #State.Fault_state := 17;
           #State.Fault_index := #State.Fault_index + 1;
         ELSIF #PBData.IW.T1_W2.Bit2 = false AND #State.Fault_index >= 0 AND #State.Fault_index <= 17 AND #State.Fault_state <> 18 THEN
           #State.Fault_state := 18;
           #State.Fault_index := 0;
         ELSIF #State.Fault_index >= 0 AND #State.Fault_index <= 17 THEN
           #State.Fault_index := 0;
         ELSE
           #State.Fault_state := 0;
           #State.Fault_index := 0;
         END_IF;
       END_IF;
     END_REGION

     // Telegramm aus dem Temp. Puffer in den DB kopieren, in Abhängigkeit des empfangenen Istwertelegrammes
     IF #IN_Sl_Akt AND #RetVal_SFC14 = 0 THEN // V1.2
       FOR #index := 0 TO 5 DO
         #Sicht_word[6 + #index] := #Empfangsdaten[#index]; // #DB_data.DW(12) := #Empfangsdaten[12];
       END_FOR;
     END_IF;                             // v1.2

     // Telegramme löschen
     IF NOT #IN_Sl_Akt OR (#IN_TL_KomF AND #RetVal_SFC14 <> 0) THEN
       FILL_BLK(IN := 16#0,
                COUNT := 23,
                OUT => #Sicht_Byte[23]);
     END_IF;
     // ProfiNet daten senden
     IF #IN_Sl_Akt THEN
       #RetVal_SFC15 := INT_TO_WORD(DPWR_DAT(LADDR := #IN_Adr, RECORD := #Sendedaten_BYTE));
     ELSE
       #RetVal_SFC15 := 0;
     END_IF;

   ELSE
     #State.Fault := FALSE;
     #State.Fault_state := 0;
   END_IF;
END_FUNCTION

FUNCTION "FC108_Pentan" : Void   // FC2, STL
{ S7_Optimized_Access := 'FALSE' }
VERSION : 0.1
   VAR_INPUT
      IN_With_Pentan : Bool;   // Pentan was requested?
      IN_With_2_Valves : Bool;   // Are there 2 filling valves existing?
      IN_ResetFault : Bool;   // Signal quit faults of this funktion block
      IN_FirstPLCcycle : Bool;   // First plc cycle
      IN_OPmode_Valid : Bool;   // A valid operation mode is selected
      IN_OPmode_Wekend : Bool;   // Operation mode weekend is selected
      IN_Filling_Selected : Bool;   // Button to select the filling
      IN_Filling_Start : Bool;   // Signal for filling the tank
      IN_Max_Level_Tank : Bool;   // Maximum level tank
      IN_Cycle_runs : Bool;   // The cycle is running
      IN_Timer_ExhauseSystem : Timer;   // Delay timer for the exhause system
      IN_Timer_Overlap_Valves : Timer;   // Delay timer to overlap the two filling valves
      IN_Timer_Valve1 : Timer;   // Switch off delay for filling valve 1
      IN_Timer_Valve2 : Timer;   // Switch off delay for filling valve 2
   END_VAR
   VAR_OUTPUT
      OUT_EnableComponent : Bool;   // Enable Filling tank with pentan
      OUT_FillingValve1 : Bool;   // Output for the filling valve 1
      OUT_FillingValve2 : Bool;   // Output for the filling valve 2
   END_VAR
   VAR_IN_OUT
      IO_Status : ANY;   // State of refilling
      IO_Fault : ANY;
      IO_NewFault : Bool;
      IO_FaultLevel_1 : Bool;
      IO_FaultLevel_2 : Bool;
      IO_FaultLevel_3 : Bool;
   END_VAR
   VAR_TEMP
      Temp_IO_Status : "UDT102_Pentan";
      ERROR_CODE : Int;   // Error state of systemfunction "BLKMOV" Blockmove
      AnyPointer1 : ANY;   // Pointer to copy thr array "IO_Status" and "Temp_IO_Status"
      AnyPointer2 : ANY;   // Pointer to copy thr array "IO_Status" and "Temp_IO_Status"
      Temp_IO_Fault : "UDT1810_Pentan";
   END_VAR
BEGIN

REGION Network 2: Saved data integration
         LAR1;
         L;
         LAR2;
   //
         L     W[AR2,P#0.0];  // Bytes
         T     W[AR1,P#0.0];
         L     W[AR2,P#2.0];  //Amount of bytes
         T     W[AR1,P#2.0];
         L     W[AR2,P#4.0];  //Block no,
         T     W[AR1,P#4.0];
         L     D[AR2,P#6.0];  //Startadress of datas
         T     D[AR1,P#6.0];
   //
         CALL  BLKMOV
         ( SRCBLK  := #AnyPointer1,
           RET_VAL := #ERROR_CODE,
           DSTBLK  := #Temp_IO_Status
         );
   //
         LAR1;
         L;
         LAR2;
   //
         L     W[AR2,P#0.0];  // Bytes
         T     W[AR1,P#0.0];
         L     W[AR2,P#2.0];  //Amount of bytes
         T     W[AR1,P#2.0];
         L     W[AR2,P#4.0];  //Block no,
         T     W[AR1,P#4.0];
         L     D[AR2,P#6.0];  //Startadress of datas
         T     D[AR1,P#6.0];
   //
         CALL  BLKMOV
         ( SRCBLK  := #AnyPointer2,
           RET_VAL := #ERROR_CODE,
           DSTBLK  := #Temp_IO_Fault
         );
   //
END_REGION

REGION Network 3: Check if pentan was requested
   // -----
         A     #IN_With_Pentan;
         JC    WithPentan;
   //-----
         AN    #IN_With_Pentan;
         =     #OUT_EnableComponent;
         =     #Temp_IO_Status.EnableComponentPump;
   //-----
         R     #Temp_IO_Fault.FLT_PreAlarm_Pentan;
         R     #Temp_IO_Fault.FLT_PreAlam_NitrogenTank;
         R     #Temp_IO_Fault.FLT_NitrogenTank;
         R     #Temp_IO_Fault.FLT_Supply_Nitrogen;
         R     #Temp_IO_Fault.FLT_Exhausesystem;
         R     #Temp_IO_Fault.FLT_PentanpumpNotRunning;
         R     #Temp_IO_Fault.FLT_PentamixNotReady;
         R     #Temp_IO_Fault.MES_EStop_Pentamix;
         R     #Temp_IO_Fault.FLT_Valve1_Max;
         R     #Temp_IO_Fault.FLT_Valve2_Max;
   //-----
         R     #Temp_IO_Status.Fault_Exist;
         R     #Temp_IO_Status.FaultLevel_1;
         R     #Temp_IO_Status.FaultLevel_2;
         R     #Temp_IO_Status.FaultLevel_3;
         R     #Temp_IO_Status.Message_Exist;
   //-----
         A     #Temp_IO_Status.HM_FillingValve;
         =     #OUT_FillingValve1;
         JU    Out;
   //-----
   WithPentan:NOP   0;
END_REGION

REGION Network 4: Fault handling
         A     #IN_ResetFault;
         R     #Temp_IO_Fault.FLT_PreAlarm_Pentan;
         R     #Temp_IO_Fault.FLT_PreAlam_NitrogenTank;
         R     #Temp_IO_Fault.FLT_NitrogenTank;
         R     #Temp_IO_Fault.FLT_Supply_Nitrogen;
         R     #Temp_IO_Fault.FLT_Exhausesystem;
         R     #Temp_IO_Fault.FLT_PentanpumpNotRunning;
         R     #Temp_IO_Fault.FLT_PentamixNotReady;
         R     #Temp_IO_Fault.FLT_Valve1_Max;
         R     #Temp_IO_Fault.FLT_Valve2_Max;
   //-----
   // Fault: Pre warning Pentan 20%
         AN    "E_Voralarm_Pentan";
         AN    #Temp_IO_Fault.FLT_PreAlarm_Pentan;
         S     #Temp_IO_Fault.FLT_PreAlarm_Pentan;
         S     #IO_FaultLevel_3;
   //-----
   // Fault: Pre warning pressure nitrogen at tank
         AN    "P_Voralarm_Stickstoff";
         AN    #Temp_IO_Fault.FLT_PreAlam_NitrogenTank;
         S     #Temp_IO_Fault.FLT_PreAlam_NitrogenTank;
         S     #IO_FaultLevel_3;
   //-----
   // Fault: Alarm nitrogen
         AN    "P_Alarm_Stickstoff";
         AN    #Temp_IO_Fault.FLT_NitrogenTank;
         S     #Temp_IO_Fault.FLT_NitrogenTank;
         S     #IO_FaultLevel_1;
   //-----
   // Fault: Supply nitrogen
         AN    "P_Alarm_VersorgungN";
         AN    #Temp_IO_Fault.FLT_Supply_Nitrogen;
         S     #Temp_IO_Fault.FLT_Supply_Nitrogen;
         S     #IO_FaultLevel_3;
   //-----
   // Fault Exhause syswtem not running
         A     #IN_OPmode_Valid;
         AN    #IN_OPmode_Wekend;
         AN    #Temp_IO_Fault.FLT_Exhausesystem;
         L     S5T#30S;
         SD    #IN_Timer_ExhauseSystem;
         A     #IN_Timer_ExhauseSystem;
         AN    "E_Absaugung_bereit";
         AN    #Temp_IO_Fault.FLT_Exhausesystem;
         S     #Temp_IO_Fault.FLT_Exhausesystem;
         S     #IO_FaultLevel_2;
   //-----
   // Message: Pentan pump not running
         A     #IN_Filling_Start;
         AN    "E_Pentanpumpe_laeuft";
         CLR;
         =     #Temp_IO_Fault.FLT_PentanpumpNotRunning;
   //-----
   // Fault: Pentamix not ready
         A     #IN_Filling_Selected;
         AN    "E_Pentamix_Ready";
         A     #IN_OPmode_Valid;
         AN    #Temp_IO_Fault.FLT_PentamixNotReady;
         CLR;
         S     #Temp_IO_Fault.FLT_PentamixNotReady;
         S     #IO_FaultLevel_3;
   //-----
   // Message: Emergecy stop from Pentamix is activ
         AN    "ES_Pentamix";
         CLR;
         =     #Temp_IO_Fault.MES_EStop_Pentamix;
   //-----
END_REGION

REGION Network 5: Enable componet with pentan
   // -----
         AN    #Temp_IO_Fault.FLT_NitrogenTank;
         =     #OUT_EnableComponent;
   //-----
         A(;
         A(;
         O     #IN_Timer_ExhauseSystem;
         O     "E_Absaugung_bereit";
         );
         AN    #Temp_IO_Fault.FLT_Exhausesystem;
         O;
         A     #IN_Cycle_runs;
         A     #Temp_IO_Fault.FLT_Exhausesystem;
         O;
         A     #IN_OPmode_Wekend;
         A     "E_Absaugung_bereit";
         );
         =     #Temp_IO_Status.EnableComponentPump;
   //-----
END_REGION

REGION Network 6: Only 1 filling valve
         A     #IN_With_2_Valves;
         JC    TwoValves;
   //-----
         AN    #IN_With_2_Valves;
         R     #Temp_IO_Status.V_FillingValve1;
         R     #Temp_IO_Status.V_FillingValve2;
         R     #OUT_FillingValve2;
         R     #Temp_IO_Fault.FLT_Valve1_Max;
         R     #Temp_IO_Fault.FLT_Valve2_Max;
   //-----
         A     #Temp_IO_Status.HM_FillingValve;
         =     #OUT_FillingValve1;
   //-----
         JU    Out;
END_REGION

REGION Network 7: Reset some signal after plc start
   TwoValves:NOP   0;
   //-----
         A     #IN_FirstPLCcycle;
         R     #Temp_IO_Status.HM_FillingValve1;
         R     #Temp_IO_Status.HM_FillingValve2;
         R     #Temp_IO_Status.HM_Valve1_closed;
         R     #Temp_IO_Status.HM_Valve2_closed;
   //-----
END_REGION
